
                       ELSE
                         // Error not matching stack type 
                         #statStatus := #ERR_PARSING;
                         #statStateIntern := #STATE_ERROR;
                         #statErrorString := CONCAT(IN1 := #statErrorString, IN2 := 'Error: No matching ');
                         #statErrorString := CONCAT(IN1 := #statErrorString, IN2 := #statKeyToken.tokenFor);
                         #statErrorString := CONCAT(IN1 := #statErrorString, IN2 := ' found to ');
                         #statErrorString := CONCAT(IN1 := #statErrorString, IN2 := #statKeyToken.tokenEndFor);
                         #statErrorString := CONCAT(IN1 := #statErrorString, IN2 := ' in line: ');
                         #statErrorString := CONCAT(IN1 := #statErrorString, IN2 := UDINT_TO_STRING(#statTokenizedLine.lineNo));
                       END_IF;
                     ELSE
                       // Error no more elements on stack
                       #statStatus := #ERR_PARSING;
                       #statStateIntern := #STATE_ERROR;
                       #statErrorString := CONCAT(IN1 := #statErrorString, IN2 := 'Error: ');
                       #statErrorString := CONCAT(IN1 := #statErrorString, IN2 := #statKeyToken.tokenEndFor);
                       #statErrorString := CONCAT(IN1 := #statErrorString, IN2 := ' not allowed in line: ');
                       #statErrorString := CONCAT(IN1 := #statErrorString, IN2 := UDINT_TO_STRING(#statTokenizedLine.lineNo));
                     END_IF;
                   END_REGION ENDFOR
                 ELSE
                   // Parse line token 
                   // Set init state for parsing line token
                   //#statStateIntern := #STATE_INIT_PARSE_LOOP;
                   #statStateIntern := #STATE_IS_LINE_SUB;
                 END_IF;

               END_IF;
             END_REGION IS_LINE_FOR

             // ------------------------------------------------------------------------------------------
             // Is line SUB
             // Check if the line contains CALL / SUB / END / M17
             // If yes then call or leave subprogram 
             // YES: Go to STATE_LINE_PARSED
             // NO: Go to PARSE_LINE_TOKENS 
             // ------------------------------------------------------------------------------------------ 
             REGION IS_LINE_SUB
               IF #statStateIntern = #STATE_IS_LINE_SUB THEN
                 // Check if line starts with 'CALL'
                 IF #statTokenizedLine.lineToken[#statTokenizedLine.numberOfToken] = #statKeyToken.tokenCallSub THEN
                   REGION CALL
                     IF #statTokenizedLine.numberOfToken >= 3 THEN // Must at least have 3 token (see below)
                       // Definition GOTO:
                       // [1] "mySub"
                       // [2] " "
                       // [3] "CALL"
                       IF #statTokenizedLine.lineToken[#statTokenizedLine.numberOfToken - 1] = ' ' // second token must be space
                         AND NOT "LKinLang_IsTokenNumberInclSign"(#statTokenizedLine.lineToken[#statTokenizedLine.numberOfToken - 2]) // labelName must not be a number
                       THEN
                         // correct jump definition 
                         // Check labelList if label exists
                         #tempLabelExists := FALSE;
                         FOR #tempLabelIndex := 1 TO #statSubPrgList.numberOfSubPrgs DO
                           IF #statSubPrgList.subPrgs[#tempLabelIndex].prgName = #statTokenizedLine.lineToken[#statTokenizedLine.numberOfToken - 2] THEN
                             // Label exists!
                             // Exit this loop
                             #tempLabelExists := TRUE;
                             EXIT;
                           END_IF;
                         END_FOR;

                         IF #tempLabelExists THEN
                           // Check if entry already exists on stack --> Avoid recursive call 
                           FOR #tempCounter := 1 TO #statStack.numberOfElements DO
                             IF #statStack.stackElements[#tempCounter].type = "LKINLANG_ENTRY_TYPE_SUB"
                               AND #statStack.stackElements[#tempCounter].quantity = #tempLabelIndex // Quantity is SubPrg index
                             THEN
                               // Sub was already called --> Error
                               #statStatus := #ERR_PARSING;
                               #statStateIntern := #STATE_ERROR;
                               #statErrorString := CONCAT(IN1 := #statErrorString, IN2 := 'Error: Recursive call of subprogram not allowed');
                               #statErrorString := CONCAT(IN1 := #statErrorString, IN2 := ' in line: ');
                               #statErrorString := CONCAT(IN1 := #statErrorString, IN2 := UDINT_TO_STRING(#statTokenizedLine.lineNo));
                               EXIT;
                             END_IF;
                           END_FOR;

                           // Check if no error occured
                           IF #statStateIntern <> #STATE_ERROR THEN
                             // Write stack entry
                             #statStack.numberOfElements += 1;
                             IF #statStack.numberOfElements <= "LKINLANG_NUMBER_OF_STACK_ELEMENTS" THEN
                               #statStack.stackElements[#statStack.numberOfElements].type := "LKINLANG_ENTRY_TYPE_SUB";
                               #statStack.stackElements[#statStack.numberOfElements].lineNumberStart := #statTokenizedLine.lineNo;
                               #statStack.stackElements[#statStack.numberOfElements].lineNumberEnd := #statSubPrgList.subPrgs[#tempLabelIndex].lineNumberEnd;
                               #statStack.stackElements[#statStack.numberOfElements].quantity := #tempLabelIndex; // Store SubPrg index as quantity
                             ELSE
                               // Error Stack overflow
                               #statStatus := #ERR_PARSING;
                               #statStateIntern := #STATE_ERROR;
                               #statErrorString := CONCAT(IN1 := #statErrorString, IN2 := 'Error: Maximum array index of stack reached');
                               #statErrorString := CONCAT(IN1 := #statErrorString, IN2 := ' in line: ');
                               #statErrorString := CONCAT(IN1 := #statErrorString, IN2 := UDINT_TO_STRING(#statTokenizedLine.lineNo));
                             END_IF;

                             // Goto line after called SUB
                             #statSearchedLine := #statSubPrgList.subPrgs[#tempLabelIndex].lineNumberStart + 1;
                             #statStateIntern := #STATE_LINE_PARSED;
                           END_IF;
                         ELSE
                           // Error: Program does not exist
                           #statStatus := #ERR_PARSING;
                           #statStateIntern := #STATE_ERROR;
                           #statErrorString := CONCAT(IN1 := #statErrorString, IN2 := 'Error: Called subprogram not found');
                           #statErrorString := CONCAT(IN1 := #statErrorString, IN2 := ' in line: ');
                           #statErrorString := CONCAT(IN1 := #statErrorString, IN2 := UDINT_TO_STRING(#statTokenizedLine.lineNo));
                         END_IF;

                       ELSE
                         // Not a correct call
                         // Throw error
                         #statStatus := #ERR_PARSING;
                         #statStateIntern := #STATE_ERROR;
                         #statErrorString := CONCAT(IN1 := #statErrorString, IN2 := 'Error: Invalid call of subprogram');
                         #statErrorString := CONCAT(IN1 := #statErrorString, IN2 := ' in line: ');
                         #statErrorString := CONCAT(IN1 := #statErrorString, IN2 := UDINT_TO_STRING(#statTokenizedLine.lineNo));
                       END_IF;
                     ELSE
                       // Not a correct call
                       // Throw error
                       #statStatus := #ERR_PARSING;
                       #statStateIntern := #STATE_ERROR;
                       #statErrorString := CONCAT(IN1 := #statErrorString, IN2 := 'Error: Invalid call of subprogram');
                       #statErrorString := CONCAT(IN1 := #statErrorString, IN2 := ' in line: ');
                       #statErrorString := CONCAT(IN1 := #statErrorString, IN2 := UDINT_TO_STRING(#statTokenizedLine.lineNo));
                     END_IF;
                   END_REGION CALL

                   // Check if line starts with 'RETURN'
                 ELSIF #statTokenizedLine.lineToken[#statTokenizedLine.numberOfToken] = #statKeyToken.tokenReturnSub THEN
                   REGION RETURN
                     IF #statTokenizedLine.numberOfToken = 1 THEN
                       IF #statStack.numberOfElements > 0 THEN
                         IF #statStack.stackElements[#statStack.numberOfElements].type = "LKINLANG_ENTRY_TYPE_SUB" THEN
                           // Goto back to line after "CALL"
                           #statSearchedLine := #statStack.stackElements[#statStack.numberOfElements].lineNumberStart + 1;
                           #statStateIntern := #STATE_LINE_PARSED;

                           // This is our scope 
                           #tempConditionCounter := DINT_TO_INT(#statStack.stackElements[#statStack.numberOfElements].quantity) * 10;

                           FOR #tempCounter := #statVarRefList.numberOfReferences TO 1 BY -1 DO
                             IF #statVarRefList.references[#tempCounter].scope = #tempConditionCounter THEN
                               // Delete variable
                               CASE #statVarRefList.references[#tempCounter].type OF
                                 "LKINLANG_VAR_TYPE_LOCAL_BOOL":
                                   #statVariables.boolean[#statVarRefList.references[#tempCounter].index] := FALSE;
                                   #statVariables.boolCounter -= 1;
                                 "LKINLANG_VAR_TYPE_LOCAL_DINT":
                                   #statVariables.dints[#statVarRefList.references[#tempCounter].index] := 0;
                                   #statVariables.dintCounter -= 1;
                                 "LKINLANG_VAR_TYPE_LOCAL_LREAL":
                                   #statVariables.lreals[#statVarRefList.references[#tempCounter].index] := 0.0;
                                   #statVariables.lrealCounter -= 1;
                               END_CASE;

                               // Delete variable reference from list
                               #statVarRefList.references[#tempCounter].index := 0;
                               #statVarRefList.references[#tempCounter].type := 0;
                               #statVarRefList.references[#tempCounter].name := '';
                               #statVarRefList.references[#tempCounter].scope := 0;
                               #statVarRefList.numberOfReferences -= 1; // Reduce number of refs
                             ELSE
                               CONTINUE;
                             END_IF;
                           END_FOR;

                           // Delete stack entry
                           #statStack.stackElements[#statStack.numberOfElements].type := 0;
                           #statStack.stackElements[#statStack.numberOfElements].lineNumberStart := 0;
                           #statStack.stackElements[#statStack.numberOfElements].lineNumberEnd := 0;
                           #statStack.stackElements[#statStack.numberOfElements].quantity := 0;
                           #statStack.numberOfElements -= 1;
                         ELSE
                           // Error not matching stack type 
                           #statStatus := #ERR_PARSING;
                           #statStateIntern := #STATE_ERROR;
                           #statErrorString := CONCAT(IN1 := #statErrorString, IN2 := 'Error: No matching ');
                           #statErrorString := CONCAT(IN1 := #statErrorString, IN2 := #statKeyToken.tokenCallSub);
                           #statErrorString := CONCAT(IN1 := #statErrorString, IN2 := ' found to ');
                           #statErrorString := CONCAT(IN1 := #statErrorString, IN2 := #statKeyToken.tokenReturnSub);
                           #statErrorString := CONCAT(IN1 := #statErrorString, IN2 := ' in line: ');
                           #statErrorString := CONCAT(IN1 := #statErrorString, IN2 := UDINT_TO_STRING(#statTokenizedLine.lineNo));
                         END_IF;
                       ELSE
                         // Error no more elements on stack
                         #statStatus := #ERR_PARSING;
                         #statStateIntern := #STATE_ERROR;
                         #statErrorString := CONCAT(IN1 := #statErrorString, IN2 := 'Error: ');
                         #statErrorString := CONCAT(IN1 := #statErrorString, IN2 := #statKeyToken.tokenEndSub);
                         #statErrorString := CONCAT(IN1 := #statErrorString, IN2 := ' not allowed in line: ');
                         #statErrorString := CONCAT(IN1 := #statErrorString, IN2 := UDINT_TO_STRING(#statTokenizedLine.lineNo));
                       END_IF;
                     ELSE
                       // Not a correct return
                       // Throw error
                       #statStatus := #ERR_PARSING;
                       #statStateIntern := #STATE_ERROR;
                       #statErrorString := CONCAT(IN1 := #statErrorString, IN2 := 'Error: Invalid return in subprogram');
                       #statErrorString := CONCAT(IN1 := #statErrorString, IN2 := ' in line: ');
                       #statErrorString := CONCAT(IN1 := #statErrorString, IN2 := UDINT_TO_STRING(#statTokenizedLine.lineNo));
                     END_IF;
                   END_REGION RETURN


                   // Check if line contains 'SUB'
                 ELSIF #statTokenizedLine.lineToken[#statTokenizedLine.numberOfToken] = #statKeyToken.tokenStartSub THEN
                   REGION SUB
                     // Throw error if SUB is found 
                     // SUB can only be written after main program
                     // and when jumping to sub the headline is skipped
                     // --> SUB should never be found in regular parsing
                     #statStatus := #ERR_PARSING;
                     #statStateIntern := #STATE_ERROR;
                     #statErrorString := CONCAT(IN1 := #statErrorString, IN2 := 'Error: ');
                     #statErrorString := CONCAT(IN1 := #statErrorString, IN2 := #statKeyToken.tokenStartSub);
                     #statErrorString := CONCAT(IN1 := #statErrorString, IN2 := ' not allowed ');
                     #statErrorString := CONCAT(IN1 := #statErrorString, IN2 := ' in line: ');
                     #statErrorString := CONCAT(IN1 := #statErrorString, IN2 := UDINT_TO_STRING(#statTokenizedLine.lineNo));
                   END_REGION SUB

                   // Check if line contains 'END / M17'
                 ELSIF FIND(IN1 := #lineBuffer.lines[#lineBuffer.pointers.retrievePointer].content, IN2 := #statKeyToken.tokenEndSub) <> 0 THEN
                   REGION END
                     IF #statTokenizedLine.numberOfToken = 2 THEN
                       IF CONCAT(IN1 := #statTokenizedLine.lineToken[#statTokenizedLine.numberOfToken], IN2 := #statTokenizedLine.lineToken[#statTokenizedLine.numberOfToken - 1]) <> #statKeyToken.tokenEndSub THEN
                         // Throw error
                         #statStatus := #ERR_PARSING;
                         #statStateIntern := #STATE_ERROR;
                         #statErrorString := CONCAT(IN1 := #statErrorString, IN2 := ';Error: Invalid end of subprogram definition');
                         #statErrorString := CONCAT(IN1 := #statErrorString, IN2 := ' in line: ');
                         #statErrorString := CONCAT(IN1 := #statErrorString, IN2 := UDINT_TO_STRING(#statTokenizedLine.lineNo));
                         EXIT;
                       END_IF;
                     ELSIF #statTokenizedLine.numberOfToken = 1 THEN
                       IF #statTokenizedLine.lineToken[#statTokenizedLine.numberOfToken] <> #statKeyToken.tokenEndSub THEN
                         // Throw error
                         #statStatus := #ERR_PARSING;
                         #statStateIntern := #STATE_ERROR;
                         #statErrorString := CONCAT(IN1 := #statErrorString, IN2 := ';Error: Invalid end of subprogram definition');
                         #statErrorString := CONCAT(IN1 := #statErrorString, IN2 := ' in line: ');
                         #statErrorString := CONCAT(IN1 := #statErrorString, IN2 := UDINT_TO_STRING(#statTokenizedLine.lineNo));
                         EXIT;
                       END_IF;
                     ELSE
                       // Throw error
                       #statStatus := #ERR_PARSING;
                       #statStateIntern := #STATE_ERROR;
                       #statErrorString := CONCAT(IN1 := #statErrorString, IN2 := ';Error: Invalid end of subprogram definition');
                       #statErrorString := CONCAT(IN1 := #statErrorString, IN2 := ' in line: ');
                       #statErrorString := CONCAT(IN1 := #statErrorString, IN2 := UDINT_TO_STRING(#statTokenizedLine.lineNo));
                       EXIT;
                     END_IF;

                     IF #statStack.numberOfElements > 0 THEN
                       IF #statStack.stackElements[#statStack.numberOfElements].type = "LKINLANG_ENTRY_TYPE_SUB" THEN
                         // Goto line after "CALL"
                         #statSearchedLine := #statStack.stackElements[#statStack.numberOfElements].lineNumberStart + 1;
                         #statStateIntern := #STATE_LINE_PARSED;

                         // This is our scope 
                         #tempConditionCounter := DINT_TO_INT(#statStack.stackElements[#statStack.numberOfElements].quantity) * 10;

                         FOR #tempCounter := #statVarRefList.numberOfReferences TO 1 BY -1 DO
                           IF #statVarRefList.references[#tempCounter].scope = #tempConditionCounter THEN
                             // Delete variable
                             CASE #statVarRefList.references[#tempCounter].type OF
                               "LKINLANG_VAR_TYPE_LOCAL_BOOL":
                                 #statVariables.boolean[#statVarRefList.references[#tempCounter].index] := FALSE;
                                 #statVariables.boolCounter -= 1;
                               "LKINLANG_VAR_TYPE_LOCAL_DINT":
                                 #statVariables.dints[#statVarRefList.references[#tempCounter].index] := 0;
                                 #statVariables.dintCounter -= 1;
                               "LKINLANG_VAR_TYPE_LOCAL_LREAL":
                                 #statVariables.lreals[#statVarRefList.references[#tempCounter].index] := 0.0;
                                 #statVariables.lrealCounter -= 1;
                             END_CASE;

                             // Delete variable reference from list
                             #statVarRefList.references[#tempCounter].index := 0;
                             #statVarRefList.references[#tempCounter].type := 0;
                             #statVarRefList.references[#tempCounter].name := '';
                             #statVarRefList.references[#tempCounter].scope := 0;
                             #statVarRefList.numberOfReferences -= 1; // Reduce number of refs
                           ELSE
                             CONTINUE;
                           END_IF;
                         END_FOR;

                         // Delete stack entry
                         #statStack.stackElements[#statStack.numberOfElements].type := 0;
                         #statStack.stackElements[#statStack.numberOfElements].lineNumberStart := 0;
                         #statStack.stackElements[#statStack.numberOfElements].lineNumberEnd := 0;
                         #statStack.stackElements[#statStack.numberOfElements].quantity := 0;
                         #statStack.numberOfElements -= 1;
                       ELSE
                         // Error not matching stack type 
                         #statStatus := #ERR_PARSING;
                         #statStateIntern := #STATE_ERROR;
                         #statErrorString := CONCAT(IN1 := #statErrorString, IN2 := 'Error: No matching ');
                         #statErrorString := CONCAT(IN1 := #statErrorString, IN2 := #statKeyToken.tokenStartSub);
                         #statErrorString := CONCAT(IN1 := #statErrorString, IN2 := ' found to ');
                         #statErrorString := CONCAT(IN1 := #statErrorString, IN2 := #statKeyToken.tokenEndSub);
                         #statErrorString := CONCAT(IN1 := #statErrorString, IN2 := ' in line: ');
                         #statErrorString := CONCAT(IN1 := #statErrorString, IN2 := UDINT_TO_STRING(#statTokenizedLine.lineNo));
                       END_IF;
                     ELSE
                       // Error no more elements on stack
                       #statStatus := #ERR_PARSING;
                       #statStateIntern := #STATE_ERROR;
                       #statErrorString := CONCAT(IN1 := #statErrorString, IN2 := 'Error: ');
                       #statErrorString := CONCAT(IN1 := #statErrorString, IN2 := #statKeyToken.tokenEndSub);
                       #statErrorString := CONCAT(IN1 := #statErrorString, IN2 := ' not allowed in line: ');
                       #statErrorString := CONCAT(IN1 := #statErrorString, IN2 := UDINT_TO_STRING(#statTokenizedLine.lineNo));
                     END_IF;
                   END_REGION END

                 ELSE
                   // Parse line token 
                   // Set init state for parsing line token
                   #statStateIntern := #STATE_INIT_PARSE_LOOP;
                 END_IF;
               END_IF;

             END_REGION IS_LINE_SUB




             // ------------------------------------------------------------------------------------------
             // Parse single tokens
             // Take one token of tokenized line and parse it
             // Use a loop to iterate over all tokens in one line
             // Go to STATE_LINE_PARSED state if all tokens are processed else keep the loop running
             // ------------------------------------------------------------------------------------------ 
             REGION PARSE_LINE_TOKEN
               // This loop is not part of a state!
               // The WHILE loop is not called if numberOfToken is 0
               // 
               // Iterate over all token in one line
               WHILE #tempTokenCounter <= #statTokenizedLine.numberOfToken
                 AND (#statStateIntern >= #STATE_INIT_PARSE_LOOP AND #statStateIntern < #STATE_LINE_PARSED)
               DO

                 // ------------------------------------------------------------------------------------------
                 // Init parse loop
                 // Initial state for one loop
                 // Initialize variables for parsing one token
                 // Next state: IS_TOKEN_SEPARATOR
                 // ------------------------------------------------------------------------------------------ 
                 REGION INIT_PARSE_LOOP
                   IF #statStateIntern = #STATE_INIT_PARSE_LOOP
                   THEN
                     // Init variables for each loop
                     #statTokenCheck.actual := #statTokenizedLine.lineToken[#tempTokenCounter];

                     // Get previous token
                     IF #tempTokenCounter > 1 THEN
                       #statTokenCheck.previous := #statTokenizedLine.lineToken[#tempTokenCounter - 1];
                     ELSE
                       #statTokenCheck.previous := '';
                     END_IF;

                     // Init parameterValid
                     #statParameterValid := #statParameterValidEmpty;

                     #statStateIntern := #STATE_IS_TOKEN_SEPARATOR;
                   END_IF;
                 END_REGION INIT_PARSE_LOOP

                 // ------------------------------------------------------------------------------------------
                 // Is token separator ?
                 // Check if token is a separator 
                 // Yes: Go to TOKEN_IS_SEPARATOR
                 // No: Go to IS_TOKEN_NUMBER
                 // ------------------------------------------------------------------------------------------ 
                 REGION IS_TOKEN_SEPARATOR
                   IF #statStateIntern = #STATE_IS_TOKEN_SEPARATOR
                   THEN
                     // Pre check if token can be separator --> Can not be if longer than 1 or is letter
                     IF LEN(#statTokenCheck.actual) > 1
                       OR "LKinLang_CharacterIsLetter"(STRING_TO_CHAR(#statTokenCheck.actual[1]))
                     THEN
                       #tempSeparatorIndex := 0;
                     ELSE
                       #tempSeparatorIndex := "LKinLang_IsTokenSeparator"(tokenToCheck := #statTokenCheck.actual, separators := #statSeparators);
                     END_IF;

                     // Decide where to go next
                     IF #tempSeparatorIndex = 0 THEN
                       #statStateIntern := #STATE_IS_TOKEN_NUMBER;
                     ELSE
                       #statStateIntern := #STATE_TOKEN_IS_SEPARATOR;
                     END_IF;
                   END_IF;
                 END_REGION IS_TOKEN_SEPARATOR

                 // ------------------------------------------------------------------------------------------
                 // Token is separator
                 // Add token to string expression if necessary
                 // Always go to TOKEN_PROCESSED
                 // ------------------------------------------------------------------------------------------ 
                 REGION TOKEN_IS_SEPARATOR
                   IF #statStateIntern = #STATE_TOKEN_IS_SEPARATOR
                   THEN
                     // Token is a separator
                     // Check if actual token is not space or equal sign --> Copy to StringExpression (e.g. math expressions)
                     IF #statTokenCheck.actual <> '=' AND #statTokenCheck.actual <> ' ' THEN
                       #statStringExpression := CONCAT(IN1 := #statTokenCheck.actual, IN2 := #statStringExpression);
                     ELSIF #statTokenCheck.actual = '=' THEN // Token is equal sign --> Change side of equation to left
                       #statRightSideOfEquation := FALSE;
                     ELSE
                       ; // Do not copy "=" & "space"  into string expression
                     END_IF;

                     #statStateIntern := #STATE_TOKEN_PROCESSED;
                   END_IF;
                 END_REGION TOKEN_IS_SEPARATOR

                 // ------------------------------------------------------------------------------------------
                 // Is token number ?
                 // Check if token is a single number 
                 // Yes: Go to TOKEN_PROCESSED
                 // No: Go to IS_TOKEN_PARAMETER
                 // ------------------------------------------------------------------------------------------ 
                 REGION IS_TOKEN_NUMBER
                   IF #statStateIntern = #STATE_IS_TOKEN_NUMBER
                   THEN
                     IF "LKinLang_IsTokenNumberInclSign"(#statTokenCheck.actual) THEN
                       IF NOT "LKinLang_CharacterIsNumeric"(#statStringExpression[1]) OR NOT #statRightSideOfEquation THEN // Check if current stringExpression contains a number
                         // Not a number --> OK
                         #statStringExpression := CONCAT(IN1 := #statTokenCheck.actual, IN2 := #statStringExpression);
                         #statStateIntern := #STATE_TOKEN_PROCESSED;
                       ELSE
                         // First char is a number --> Cannot concat two numbers in a row --> ERROR
                         #statStatus := #ERR_PARSING;
                         #statErrorString := CONCAT(IN1 := #statErrorString, IN2 := 'Error: Invalid syntax');
                         #statErrorString := CONCAT(IN1 := #statErrorString, IN2 := '; Line: ');
                         #statErrorString := CONCAT(IN1 := #statErrorString, IN2 := UDINT_TO_STRING(#statTokenizedLine.lineNo));
                         EXIT;
                       END_IF;
                     ELSE
                       #statStateIntern := #STATE_IS_TOKEN_PARAMETER;
                     END_IF;
                   END_IF;
                 END_REGION IS_TOKEN_NUMBER

                 // ------------------------------------------------------------------------------------------
                 // Is token parameter
                 // Check if token is parameter defined in the selected language
                 // YES: Go to TOKEN_IS_PARAMETER 
                 // NO: Go to IS_TOKEN_VARIABLE
                 // ------------------------------------------------------------------------------------------ 
                 REGION IS_TOKEN_PARAMETER
                   IF #statStateIntern = #STATE_IS_TOKEN_PARAMETER
                   THEN
                     // Reset parameter definition
                     #statParameterDefinition := #statParameterDefinitionEmpty;

                     // Check if Token is parameter 
                     #tempParameterIndex := "LKinLang_IsTokenParameter"(tokenToCheck := #statTokenCheck,
                                                                        language := #language,
                                                                        lastIndexLookUp := #statLastIndexLookUp,
                                                                        parameterDefinition := #statParameterDefinition,
                                                                        parameterLookUpTable := #statParameterLookUpTable,
                                                                        parameterDefaults := #parameterDefaults,
                                                                        directCmdWord := #statDirectCmdWord,
                                                                        configCmdWords := #statConfigCmdWords);

                     // Decide where to go next
                     IF #tempParameterIndex = 0 THEN
                       #statStateIntern := #STATE_IS_TOKEN_VARIABLE;
                     ELSE
                       #statStateIntern := #STATE_TOKEN_IS_PARAMETER;
                     END_IF;

                   END_IF;
                 END_REGION IS_TOKEN_PARAMETER

                 // ------------------------------------------------------------------------------------------
                 // Token is parameter
                 // Token was found to be a parameter in the seleceted language
                 // Definition is already found
                 // Translate into path data
                 // ------------------------------------------------------------------------------------------ 
                 REGION TOKEN_IS_PARAMETER
                   IF #statStateIntern = #STATE_TOKEN_IS_PARAMETER
                   THEN

                     // Carefull! Is this really necessary ??
                     // Delete String expression if parameter has a number (like G01, ...)
                     IF #statParameterDefinition.parameterNameNumber <> -1
                       AND NOT "LKinLang_CheckProperty"(properties := #statParameterDefinition.properties, propertyToCheck := "LKINLANG_EQUATION")
                     THEN
                       #statStringExpression := '';
                     END_IF;

                     REGION SET_CONDITIONS
                       // Set parameter in found conditions arrays and also get conditions to check from parameter
                       "LKinLang_SetParameterConditions"(parameterNumber := #tempParameterIndex,
                                                         tempParameterDef := #statParameterDefinition,
                                                         parametersInLine := #statSetParametersInLine,
                                                         parametersInCommand := #statSetParametersInCmd,
                                                         parametersInProgram := #statSetParametersInPrg,
                                                         conditionsToCheck := #statConditionsToCheck,
                                                         conditionCounter := #tempConditionCounter);
                     END_REGION SET_CONDITIONS

                     REGION CHECK_PARAMETER_COUNTER
                       // Check if same parameter was set more than validCountsPerLine
                       "LKinLang_CheckParameterCounter"(parameterNumber := #tempParameterIndex,
                                                        parameterDefinition := #statParameterDefinition,
                                                        lineNo := #statTokenizedLine.lineNo,
                                                        parameterCounter := #tempParameterCounter,
                                                        errorString := #statErrorString,
                                                        error := #tempError);

                       IF #tempError THEN
                         #statStatus := #ERR_PARSING;
                         // error string is alread written
                         EXIT;
                       END_IF;
                     END_REGION CHECK_PARAMETER_COUNTER

                     REGION CHECK_PROPERTIES
                       // Check for motion command
                       IF "LKinLang_CheckProperty"(properties := #statParameterDefinition.properties, propertyToCheck := "LKINLANG_MOTION_CMD") THEN
                         #statModalCommand.motionCmd := #tempParameterIndex;
                       END_IF;

                       // Copy properties to actual command
                       #statActualCommand.properties := #statParameterDefinition.properties;

                       // Check for relative or absolute positioning property
                       IF
                         "LKinLang_CheckProperty"(properties := #statParameterDefinition.properties, propertyToCheck := "LKINLANG_ABSOLUTE_POSITION")
                         AND
                         "LKinLang_CheckProperty"(properties := #statParameterDefinition.properties, propertyToCheck := "LKINLANG_RELATIVE_POSITION")
                       THEN
                         #statStatus := #ERR_PARSING;
                         #statErrorString := 'Error: Position setting invalid';
                         #statErrorString := CONCAT(IN1 := #statErrorString, IN2 := '; Line: ');
                         #statErrorString := CONCAT(IN1 := #statErrorString, IN2 := UDINT_TO_STRING(#statTokenizedLine.lineNo));
                         EXIT;

                       ELSIF "LKinLang_CheckProperty"(properties := #statParameterDefinition.properties, propertyToCheck := "LKINLANG_RELATIVE_POSITION") THEN
                         #statPositioningMode := 2; // Relative positions

                       ELSIF "LKinLang_CheckProperty"(properties := #statParameterDefinition.properties, propertyToCheck := "LKINLANG_ABSOLUTE_POSITION") THEN
                         #statPositioningMode := 1; // Absolute positions

                       ELSE
                         ; // No position property set --> do nothing
                       END_IF;

                     END_REGION CHECK_PROPERTIES


                     // ------------------------------------------------------------------------------------------
                     // Translate to pathdata
                     //
                     // Maybe check Prio of actual parsed cmd and then set if same or higher ?
                     // Do Priority check from FC SetVal before calling set val as it is not usefull to check all things and then cancel because of prio
                     // 
                     // Something like this 
                     // 1. Parse/get the Follow values into separate variable
                     // 2. Call FC SetValue for each follow value where necessary
                     // 3. Parse the direct values --> Check if priority was already written in step 2
                     // --> Only write if priority is higher (in one parameter one variable can only have one prio for follow val and direct val)
                     // --> each path data var will have direct val and follow val with same prio 
                     // --> Generate no error message when same prio
                     // 
                     // IF #actualCommand.priority < statParameterDef.priorities then 
                     //    FC SetVal
                     // ELSE
                     //    parameter was set with same or higher prio   
                     // END_IF
                     // ------------------------------------------------------------------------------------------
                     // 
                     // First run: Get follow values and write path data element
                     // Second run: Get direct values and write path data element
                     FOR #tempParseCounter := 1 TO 2 DO

                       IF #tempParseCounter = 1 THEN
                         REGION GET_FOLLOW_VALUES
                           // Copy CmdWords to temp
                           FOR #tempFollowValueCounter := 1 TO "LKINLANG_NUMBER_OF_FOLLOW_VALUES" DO
                             #tempCmdWord := #tempCmdWord OR #statConfigCmdWords[#tempFollowValueCounter];
                           END_FOR;

                           // Config Commands check and set the programmed value after the parameter (e.g. F200)
                           // Check if follow value are to be set
                           FOR #tempFollowValueCounter := 1 TO "LKINLANG_NUMBER_OF_FOLLOW_VALUES" DO
                             IF NOT #statConfigCmdWords[#tempFollowValueCounter].%X0 // Check if at least one follow val is configured
                               OR #statStringExpression = ''
                             THEN
                               EXIT;
                             ELSE
                               // Add exception when parsing H Parameter 
                               // G1 X100 H100=12.3 
                               // OR
                               // G1 X100 H100 = 12.3
                               // Problem: "=" is not added to StringExpression
                               // --> GetValue is not working correctly as more follow values have to be separated by ","
                               //
                               // StringExpression looks like:
                               // "10012.3"
                               // only rigthSideOfEquation=false indicates that a "=" was there
                               // 
                               // Check string expression and add "," if necessary
                               IF #statRightSideOfEquation = FALSE AND #tempFollowValueCounter = 1 THEN
                                 // Search right place in stringExpression and add a "," ?
                                 #tempCounter := FIND(IN1 := #statStringExpression, IN2 := #statTokenCheck.previous);

                                 IF #tempCounter <> 0 THEN
                                   #statStringExpression := INSERT(IN1 := #statStringExpression, IN2 := ',', P := #tempCounter + LEN(#statTokenCheck.previous) - 1);
                                 END_IF;
                               END_IF;

                               // Get parameter value
                               #tempReturnVal := "LKinLang_GetValue"(tokenNo := #tempTokenCounter,
                                                                     properties := #statParameterDefinition.properties,
                                                                     parameterValue => #tempParameterValue,
                                                                     followValCounter := #tempFollowValueCounter,
                                                                     stringExpression := #statStringExpression,
                                                                     errorString := #statErrorString,
                                                                     token := #statTokenizedLine);

                               IF #tempReturnVal <> 0 THEN
                                 // Error
                                 #statStatus := #ERR_PARSING;
                                 #statErrorString := CONCAT(IN1 := #statErrorString, IN2 := '; Line: ');
                                 #statErrorString := CONCAT(IN1 := #statErrorString, IN2 := UDINT_TO_STRING(#statTokenizedLine.lineNo));
                                 EXIT;
                               END_IF;


                               REGION CMD_TYPE
                                 // Command type
                                 IF #statParameterDefinition.followingValues[#tempFollowValueCounter].cmdType THEN
                                   #tempParsedValues.cmdType := LREAL_TO_INT(#tempParameterValue);
                                   #statParameterValid.cmdType := TRUE;
                                 END_IF;
                               END_REGION CMD_TYPE

                               REGION CMD_NAME  
                                 // Command name
                                 IF #statParameterDefinition.followingValues[#tempFollowValueCounter].cmdName THEN
                                   // 16.07.2019 FR: Changed conversion function and checked if string does not overflow
                                   #tempCmdName := "LKinLang_LRealToReducedString"(input := #tempParameterValue, decimalPlaces := 0);
                                   IF LEN(#tempCmdName) <= MAX_LEN(#tempParsedValues.cmdName) THEN
                                     #tempParsedValues.cmdName := #tempCmdName;
                                     #statParameterValid.cmdName := TRUE;
                                   ELSE
                                     // Error string: length not sufficient
                                     #statStatus := #ERR_PARSING;
                                     #statErrorString := CONCAT(IN1 := #statErrorString, IN2 := 'Command name too long');
                                     #statErrorString := CONCAT(IN1 := #statErrorString, IN2 := '; Line: ');
                                     #statErrorString := CONCAT(IN1 := #statErrorString, IN2 := UDINT_TO_STRING(#statTokenizedLine.lineNo));
                                     EXIT;
                                   END_IF;
                                 END_IF;
                               END_REGION CMD_NAME

                               REGION COORDINATES
                                 IF #statConfigCmdWords[#tempFollowValueCounter].%X1 THEN
                                   // X coordinate
                                   IF #statParameterDefinition.followingValues[#tempFollowValueCounter].cmdCoordinates.cartesianPosition.x THEN
                                     #tempParsedValues.cmdCoordinates.cartesianPosition.x := #tempParameterValue;
                                     #statParameterValid.cmdCoordinates.cartesianPosition.x := TRUE;
                                   END_IF;

                                   // Y coordinate
                                   IF #statParameterDefinition.followingValues[#tempFollowValueCounter].cmdCoordinates.cartesianPosition.y THEN
                                     #tempParsedValues.cmdCoordinates.cartesianPosition.y := #tempParameterValue;
                                     #statParameterValid.cmdCoordinates.cartesianPosition.y := TRUE;
                                   END_IF;

                                   // Z coordinate
                                   IF #statParameterDefinition.followingValues[#tempFollowValueCounter].cmdCoordinates.cartesianPosition.z THEN
                                     #tempParsedValues.cmdCoordinates.cartesianPosition.z := #tempParameterValue;
                                     #statParameterValid.cmdCoordinates.cartesianPosition.z := TRUE;
                                   END_IF;

                                   // A coordinate
                                   IF #statParameterDefinition.followingValues[#tempFollowValueCounter].cmdCoordinates.cartesianPosition.a THEN
                                     #tempParsedValues.cmdCoordinates.cartesianPosition.a := #tempParameterValue;
                                     #statParameterValid.cmdCoordinates.cartesianPosition.a := TRUE;
                                   END_IF;

                                   // Coordinate System
                                   IF #statParameterDefinition.followingValues[#tempFollowValueCounter].cmdCoordinates.coordSystem THEN
                                     #tempParsedValues.cmdCoordinates.coordSystem := LREAL_TO_DINT(#tempParameterValue);
                                     #statParameterValid.cmdCoordinates.coordSystem := TRUE;
                                   END_IF;
                                 END_IF;
                               END_REGION COORDINATES

                               REGION GENERAL_PARAMETERS
                                 IF #statConfigCmdWords[#tempFollowValueCounter].%X2 THEN

                                   // Buffermode
                                   IF #statParameterDefinition.followingValues[#tempFollowValueCounter].cmdParameters.bufferMode THEN
                                     // Set Buffermode
                                     #tempParsedValues.cmdParameters.bufferMode := LREAL_TO_DINT(#tempParameterValue);
                                     #statParameterValid.cmdParameters.bufferMode := TRUE;
                                   END_IF;


                                   // DynamicAdaption
                                   IF #statParameterDefinition.followingValues[#tempFollowValueCounter].cmdParameters.dynamicAdaption THEN
                                     // Set DynamicAdaption
                                     #tempParsedValues.cmdParameters.dynamicAdaption := LREAL_TO_DINT(#tempParameterValue);
                                     #statParameterValid.cmdParameters.dynamicAdaption := TRUE;
                                   END_IF;

                                   // Offset Parameter
                                   // Offset ParaNo
                                   IF #statParameterDefinition.followingValues[#tempFollowValueCounter].cmdParameters.offsetParameters.offsetParaNo THEN
                                     // Set OffsetParaNo
                                     #tempParsedValues.cmdParameters.offsetParameters.offsetParaNo := LREAL_TO_INT(#tempParameterValue);
                                     #statParameterValid.cmdParameters.offsetParameters.offsetParaNo := TRUE;
                                   END_IF;

                                   // OffsetMainPathPlane
                                   IF #statParameterDefinition.followingValues[#tempFollowValueCounter].cmdParameters.offsetParameters.mainPathPlane THEN
                                     // Set Main path plane
                                     #tempParsedValues.cmdParameters.offsetParameters.mainPathPlane := LREAL_TO_INT(#tempParameterValue);
                                     #statParameterValid.cmdParameters.offsetParameters.mainPathPlane := TRUE;
                                   END_IF;

                                   // Transition parameter
                                   FOR #tempCounter := 1 TO 5 DO
                                     // Transition Parameter
                                     IF #statParameterDefinition.followingValues[#tempFollowValueCounter].cmdParameters.transitionParameters[#tempCounter] THEN
                                       // Set Transition Parameter
                                       #tempParsedValues.cmdParameters.transitionParameters[#tempCounter] := #tempParameterValue;
                                       #statParameterValid.cmdParameters.transitionParameters[#tempCounter] := TRUE;
                                     END_IF;
                                   END_FOR;

                                 END_IF;
                               END_REGION GENERAL_PARAMETERS

                               REGION PATH_DYNAMICS
                                 IF #statConfigCmdWords[#tempFollowValueCounter].%X3 THEN

                                   // Velocity
                                   IF #statParameterDefinition.followingValues[#tempFollowValueCounter].cmdParameters.pathDynamics.velocity THEN
                                     #tempParsedValues.cmdParameters.pathDynamics.velocity := #tempParameterValue;
                                     #statParameterValid.cmdParameters.pathDynamics.velocity := TRUE;
                                   END_IF;

                                   // Acceleration
                                   IF #statParameterDefinition.followingValues[#tempFollowValueCounter].cmdParameters.pathDynamics.acceleration THEN
                                     #tempParsedValues.cmdParameters.pathDynamics.acceleration := #tempParameterValue;
                                     #statParameterValid.cmdParameters.pathDynamics.acceleration := TRUE;
                                   END_IF;

                                   // Deceleration
                                   IF #statParameterDefinition.followingValues[#tempFollowValueCounter].cmdParameters.pathDynamics.deceleration THEN
                                     #tempParsedValues.cmdParameters.pathDynamics.deceleration := #tempParameterValue;
                                     #statParameterValid.cmdParameters.pathDynamics.deceleration := TRUE;
                                   END_IF;

                                   // Jerk
                                   IF #statParameterDefinition.followingValues[#tempFollowValueCounter].cmdParameters.pathDynamics.jerk THEN
                                     #tempParsedValues.cmdParameters.pathDynamics.jerk := #tempParameterValue;
                                     #statParameterValid.cmdParameters.pathDynamics.jerk := TRUE;
                                   END_IF;

